screen "1. MAIN" 1280x800, template "Main_Template"
   on GenerateScreen: SetTag("animation_page", 1)
   Softkey "Softkey_F1" at 0,0 size 0x0
      on KeyDown: ActivateScreen("1. MAIN", 0)
   Softkey "Softkey_F2" at 0,0 size 0x0
      on KeyDown: ActivateScreen("2. VFD 2 - 5", 0)
   Softkey "Softkey_F3" at 0,0 size 0x0
      on KeyDown: ActivateScreen("3. VFD 6 - 9", 0)
   Softkey "Softkey_F4" at 0,0 size 0x0
      on KeyDown: ActivateScreen("4. VFD 10 - 13", 0)
   Softkey "Softkey_F5" at 0,0 size 0x0
      on KeyDown: ActivateScreen("5. VFD 14 - 17", 0)
   Softkey "Softkey_F6" at 0,0 size 0x0
      on KeyDown: ActivateScreen("6. VFD 18 - 21", 0)
   Softkey "Softkey_F7" at 0,0 size 0x0
      on KeyDown: ActivateScreen("7. VFD 22 - 23", 0)
   Softkey "Softkey_F8" at 0,0 size 0x0
      on KeyDown: ActivateScreen("8. ALARM", 0)
   Softkey "Softkey_F9" at 0,0 size 0x0
      on KeyDown: ActivateScreen("9. VFD PROFIBUS", 0)
   Softkey "Softkey_F10" at 0,0 size 0x0
      on KeyDown: ActivateScreen("10. SETTINGS", 0)
   TextField "Text field_33" at 632,247 size 105x42; Text 'Hz'
   TextField "Text field_1" at 0,64 size 331x50; Text 'ACTUAL MOTOR SPEED'
   Button "Button_1" at 0,721 size 160x79; TextOff 'MAIN'
      on Click: ActivateScreen("1. MAIN", 0)
      Appearance <- "animation_page"
   Button "Button_10" at 160,721 size 160x79; TextOff 'VFD 2 - 5'
      on Click: ActivateScreen("2. VFD 2 - 5", 0)
      Appearance <- "animation_page"
   Button "Button_11" at 320,721 size 160x79; TextOff 'VFD 6 - 9'
      on Click: ActivateScreen("3. VFD 6 - 9", 0)
      Appearance <- "animation_page"
   Button "Button_12" at 480,721 size 160x79; TextOff 'VFD 10 - 13'
      on Click: ActivateScreen("4. VFD 10 - 13", 0)
      Appearance <- "animation_page"
   Button "Button_13" at 640,721 size 160x79; TextOff 'VFD 14 - 17'
      on Click: ActivateScreen("5. VFD 14 - 17", 0)
      Appearance <- "animation_page"
   Button "Button_14" at 800,721 size 160x79; TextOff 'VFD 18 - 21'
      on Click: ActivateScreen("6. VFD 18 - 21", 0)
      Appearance <- "animation_page"
   Button "Button_15" at 960,721 size 160x79; TextOff 'VFD 22 - 23'
      on Click: ActivateScreen("7. VFD 22 - 23", 0)
      Appearance <- "animation_page"
   Button "Button_16" at 1120,721 size 160x79; TextOff 'Alarm'
      on Click: ActivateScreen("8. ALARM", 0)
      Appearance <- "animation_page"
   Group "Group" at 90,528 size 42x28
   Group "Group_1" at 57,540 size 42x28
   Group "Group_4" at 657,193 size 42x28
   Group "Group_5" at 3,194 size 42x28
   Group "Group_6" at 41,515 size 42x28
   Group "Group_15" at 926,512 size 42x28
   Group "Group_16" at 1063,535 size 42x28
   Group "Group_17" at 1008,534 size 42x28
   Group "Group_19" at 1058,421 size 42x28
   Group "Group_20" at 1103,421 size 42x28
   Group "Group_21" at 1165,505 size 42x28
   Group "Group_10" at 547,540 size 42x28
   Group "Group_9" at 510,515 size 42x28
   Group "Group_7" at 358,515 size 42x28
   Group "Group_8" at 396,540 size 42x28
   Group "Group_2" at 210,515 size 42x28
   Group "Group_3" at 252,540 size 42x28
   Group "Group_11" at 660,540 size 42x28
   Group "Group_12" at 797,502 size 42x28
   Group "Group_13" at 797,540 size 42x28
   Group "Group_14" at 853,530 size 42x28
   IOField "I/O field_17" at 633,252 size 60x33; FormatPattern 99.99
      ProcessValue <- "speedActual_address_18"
   TextField "Text field_24" at 22,247 size 105x42; Text 'Hz'
   IOField "I/O field_1" at 24,252 size 60x33; FormatPattern 99.99
      ProcessValue <- "speedActual_address_2"
   TextField "Text field_25" at 10,342 size 105x42; Text 'Hz'
   IOField "I/O field_2" at 12,347 size 60x33; FormatPattern 99.99
      ProcessValue <- "speedActual_address_3"
   Circle "Circle_34" at 693,170 size 28x28
      Appearance <- "Running_Motor Addres_23"
   Group "Group_18" at 1203,505 size 42x28
   Group "Group_22" at 1186,539 size 42x28
   Group "Group_23" at 11,162 size 42x28
   Group "Group_24" at 657,161 size 42x28
   TextField "Text field_29" at 33,653 size 105x42; Text 'Hz'
   IOField "I/O field_3" at 33,658 size 60x33; FormatPattern 99.99
      ProcessValue <- "speedActual_address_4"
   TextField "Text field_30" at 85,604 size 105x42; Text 'Hz'
   IOField "I/O field_4" at 87,609 size 60x33; FormatPattern 99.99
      ProcessValue <- "speedActual_address_5"
   TextField "Text field_31" at 177,653 size 105x42; Text 'Hz'
   IOField "I/O field_5" at 177,658 size 60x33; FormatPattern 99.99
      ProcessValue <- "speedActual_address_6"
   TextField "Text field_32" at 245,604 size 105x42; Text 'Hz'
   IOField "I/O field_6" at 247,609 size 60x33; FormatPattern 99.99
      ProcessValue <- "speedActual_address_7"
   TextField "Text field_34" at 322,653 size 105x42; Text 'Hz'
   IOField "I/O field_7" at 322,658 size 60x33; FormatPattern 99.99
      ProcessValue <- "speedActual_address_8"
   TextField "Text field_35" at 386,604 size 105x42; Text 'Hz'
   IOField "I/O field_8" at 388,609 size 60x33; FormatPattern 99.99
      ProcessValue <- "speedActual_address_9"
   TextField "Text field_36" at 467,653 size 105x42; Text 'Hz'
   IOField "I/O field_9" at 467,658 size 60x33; FormatPattern 99.99
      ProcessValue <- "speedActual_address_10"
   TextField "Text field_37" at 542,604 size 105x42; Text 'Hz'
   IOField "I/O field_10" at 544,609 size 60x33; FormatPattern 99.99
      ProcessValue <- "speedActual_address_11"
   TextField "Text field_38" at 611,653 size 105x42; Text 'Hz'
   IOField "I/O field_11" at 611,658 size 60x33; FormatPattern 99.99
      ProcessValue <- "speedActual_address_12"
   TextField "Text field_39" at 742,604 size 105x42; Text 'Hz'
   IOField "I/O field_12" at 744,609 size 60x33; FormatPattern 99.99
      ProcessValue <- "speedActual_address_13"
   TextField "Text field_40" at 756,653 size 105x42; Text 'Hz'
   IOField "I/O field_13" at 756,658 size 60x33; FormatPattern 99.99
      ProcessValue <- "speedActual_address_15"
   TextField "Text field_41" at 700,382 size 105x42; Text 'Hz'
   IOField "I/O field_14" at 702,387 size 60x33; FormatPattern 99.99
      ProcessValue <- "speedActual_address_14"
   TextField "Text field_42" at 901,653 size 105x42; Text 'Hz'
   IOField "I/O field_15" at 901,658 size 60x33; FormatPattern 99.99
      ProcessValue <- "speedActual_address_16"
   TextField "Text field_43" at 970,604 size 105x42; Text 'Hz'
   IOField "I/O field_16" at 972,609 size 60x33; FormatPattern 99.99
      ProcessValue <- "speedActual_address_17"
   TextField "Text field_44" at 1046,653 size 105x42; Text 'Hz'
   IOField "I/O field_18" at 1048,658 size 60x33; FormatPattern 99.99
      ProcessValue <- "speedActual_address_19"
   TextField "Text field_45" at 1150,604 size 105x42; Text 'Hz'
   IOField "I/O field_19" at 1152,609 size 60x33; FormatPattern 99.99
      ProcessValue <- "speedActual_address_22"
   TextField "Text field_46" at 1170,403 size 105x42; Text 'Hz'
   IOField "I/O field_20" at 1172,408 size 60x33; FormatPattern 99.99
      ProcessValue <- "speedActual_address_21"
   TextField "Text field_47" at 1170,325 size 105x42; Text 'Hz'
   IOField "I/O field_21" at 1172,330 size 60x33; FormatPattern 99.99
      ProcessValue <- "speedActual_address_20"
   TextField "Text field_48" at 1054,298 size 105x42; Text 'Hz'
   IOField "I/O field_22" at 1056,303 size 60x33; FormatPattern 99.99
      ProcessValue <- "speedActual_address_23"
   TextField "Text field_49" at 629,117 size 105x42; Text 'Hz'
   IOField "I/O field_23" at 631,122 size 60x33; FormatPattern 99.99
      ProcessValue <- "speedActual_address_23"
   TextField "Text field_50" at 13,117 size 105x42; Text 'Hz'
   IOField "I/O field_24" at 15,122 size 60x33; FormatPattern 99.99
      ProcessValue <- "speedActual_address_23"
   TextField "Text field_87" at 873,193 size 190x45; Text 'Rotary Moulder'
   Circle "Circle_10" at 883,201 size 29x29
      Appearance <- "Syncron_1"
   TextField "Text field_88" at 1071,141 size 190x45; Text 'Rotary Cutter'
   Circle "Circle_11" at 1081,149 size 29x29
      Appearance <- "Syncron_2"
   TextField "Text field_95" at 1071,193 size 190x45; Text 'Swivel Panner'
   Circle "Circle_12" at 1081,200 size 29x29
      Appearance <- "Syncron_3"
   TextField "Text field_51" at 873,141 size 190x45; Text 'SYNC MODE'
   TextField "Text field_52" at 42,320 size 42x25; Text '3'
   TextField "Text field_53" at 65,692 size 42x25; Text '4'
   TextField "Text field_54" at 117,582 size 42x25; Text '5'
   TextField "Text field_55" at 54,224 size 42x25; Text '2'
   TextField "Text field_56" at 635,224 size 42x25; Text '18'
   TextField "Text field_57" at 593,124 size 42x25; Text '23'
   TextField "Text field_58" at 121,124 size 42x25; Text '23'
   TextField "Text field_59" at 1086,276 size 42x25; Text '23'
   TextField "Text field_60" at 1173,582 size 42x25; Text '22'
   TextField "Text field_61" at 1202,300 size 42x25; Text '20'
   TextField "Text field_62" at 1202,376 size 42x25; Text '21'
   TextField "Text field_63" at 209,692 size 42x25; Text '6'
   TextField "Text field_64" at 277,582 size 42x25; Text '7'
   TextField "Text field_65" at 354,692 size 42x25; Text '8'
   TextField "Text field_66" at 418,582 size 42x25; Text '9'
   TextField "Text field_67" at 499,692 size 42x25; Text '10'
   TextField "Text field_68" at 574,582 size 42x25; Text '11'
   TextField "Text field_69" at 643,692 size 42x25; Text '12'
   TextField "Text field_70" at 788,692 size 42x25; Text '15'
   TextField "Text field_71" at 732,358 size 42x25; Text '14'
   TextField "Text field_72" at 990,582 size 42x25; Text '17'
   TextField "Text field_73" at 933,692 size 42x25; Text '16'
   TextField "Text field_74" at 1078,692 size 42x25; Text '19'
   TextField "Text field_75" at 774,582 size 42x25; Text '13'
   Button "Button_2" at 4,193 size 42x36; TextOff 'Text'
      on Click: ActivateScreen("2. VFD 2 - 5", 0)
   Button "Button_3" at 42,508 size 43x38; TextOff 'Text'
      on Click: ActivateScreen("2. VFD 2 - 5", 0)
   Button "Button_4" at 217,510 size 33x39; TextOff 'Text'
      on Click: ActivateScreen("3. VFD 6 - 9", 0)
   Button "Button_5" at 360,510 size 36x40; TextOff 'Text'
      on Click: ActivateScreen("3. VFD 6 - 9", 0)
   Button "Button_6" at 513,510 size 38x40; TextOff 'Text'
      on Click: ActivateScreen("4. VFD 10 - 13", 0)
   Button "Button_7" at 663,532 size 40x41; TextOff 'Text'
      on Click: ActivateScreen("4. VFD 10 - 13", 0)
   Button "Button_8" at 548,532 size 38x40; TextOff 'Text'
      on Click: ActivateScreen("4. VFD 10 - 13", 0)
   Button "Button_9" at 799,532 size 40x41; TextOff 'Text'
      on Click: ActivateScreen("4. VFD 10 - 13", 0)
   Button "Button_17" at 855,524 size 40x41; TextOff 'Text'
      on Click: ActivateScreen("5. VFD 14 - 17", 0)
   Button "Button_18" at 799,492 size 40x41; TextOff 'Text'
      on Click: ActivateScreen("5. VFD 14 - 17", 0)
   Button "Button_19" at 927,508 size 40x41; TextOff 'Text'
      on Click: ActivateScreen("5. VFD 14 - 17", 0)
   Button "Button_20" at 1007,524 size 40x41; TextOff 'Text'
      on Click: ActivateScreen("5. VFD 14 - 17", 0)
   Button "Button_21" at 1064,526 size 40x41; TextOff 'Text'
      on Click: ActivateScreen("6. VFD 18 - 21", 0)
   Button "Button_22" at 1187,539 size 40x31; TextOff 'Text'
      on Click: ActivateScreen("7. VFD 22 - 23", 0)
   Button "Button_23" at 1165,497 size 82x41; TextOff 'Text'
      on Click: ActivateScreen("6. VFD 18 - 21", 0)
   Button "Button_24" at 1060,414 size 40x39; TextOff 'Text'
      on Click: ActivateScreen("7. VFD 22 - 23", 0)
   Button "Button_25" at 1105,414 size 40x39; TextOff 'Text'
      on Click: ActivateScreen("7. VFD 22 - 23", 0)
   Button "Button_26" at 659,156 size 40x39; TextOff 'Text'
      on Click: ActivateScreen("7. VFD 22 - 23", 0)
   Button "Button_27" at 13,156 size 40x39; TextOff 'Text'
      on Click: ActivateScreen("7. VFD 22 - 23", 0)
   Button "Button_28" at 659,190 size 40x41; TextOff 'Text'
      on Click: ActivateScreen("6. VFD 18 - 21", 0)
   Button "Button_29" at 400,533 size 36x40; TextOff 'Text'
      on Click: ActivateScreen("3. VFD 6 - 9", 0)
   Button "Button_30" at 257,534 size 33x39; TextOff 'Text'
      on Click: ActivateScreen("3. VFD 6 - 9", 0)
   Button "Button_31" at 58,532 size 43x38; TextOff 'Text'
      on Click: ActivateScreen("2. VFD 2 - 5", 0)
   Button "Button_32" at 90,524 size 43x38; TextOff 'Text'
      on Click: ActivateScreen("2. VFD 2 - 5", 0)
   Circle "Circle_2" at 97,528 size 28x28
      Appearance <- "Running_Motor Addres_5"
   TextField "Text field_2" at 90,530 size 42x25; Text 'M'
   Circle "Circle_23" at 64,540 size 28x28
      Appearance <- "Running_Motor Addres_4"
   TextField "Text field_3" at 57,542 size 42x25; Text 'M'
   Circle "Circle_6" at 664,193 size 28x28
      Appearance <- "Running_Motor Addres_18"
   TextField "Text field_6" at 657,195 size 42x25; Text 'M'
   Circle "Circle_22" at 10,194 size 28x28
      Appearance <- "Running_Motor Addres_2"
   TextField "Text field_7" at 3,196 size 42x25; Text 'M'
   Circle "Circle_5" at 48,515 size 28x28
      Appearance <- "Running_Motor Addres_3"
   TextField "Text field_8" at 41,517 size 42x25; Text 'M'
   Circle "Circle_31" at 933,512 size 28x28
      Appearance <- "Running_Motor Addres_16"
   TextField "Text field_17" at 926,514 size 42x25; Text 'M'
   Circle "Circle_32" at 1070,535 size 28x28
      Appearance <- "Running_Motor Addres_19"
   TextField "Text field_18" at 1063,537 size 42x25; Text 'M'
   Circle "Circle_33" at 1015,534 size 28x28
      Appearance <- "Running_Motor Addres_17"
   TextField "Text field_19" at 1008,536 size 42x25; Text 'M'
   Circle "Circle_35" at 1065,421 size 28x28
      Appearance <- "Running_Motor Addres_23"
   TextField "Text field_21" at 1058,423 size 42x25; Text 'M'
   Circle "Circle_36" at 1110,421 size 28x28
      Appearance <- "Running_Motor Addres_23"
   TextField "Text field_22" at 1103,423 size 42x25; Text 'M'
   Circle "Circle_37" at 1172,505 size 28x28
      Appearance <- "Running_Motor Addres_20"
   TextField "Text field_23" at 1165,507 size 42x25; Text 'M'
   Circle "Circle_26" at 554,540 size 28x28
      Appearance <- "Running_Motor Addres_11"
   TextField "Text field_12" at 547,542 size 42x25; Text 'M'
   Circle "Circle_25" at 517,515 size 28x28
      Appearance <- "Running_Motor Addres_10"
   TextField "Text field_11" at 510,517 size 42x25; Text 'M'
   Circle "Circle_21" at 365,515 size 28x28
      Appearance <- "Running_Motor Addres_8"
   TextField "Text field_9" at 358,517 size 42x25; Text 'M'
   Circle "Circle_24" at 403,540 size 28x28
      Appearance <- "Running_Motor Addres_9"
   TextField "Text field_10" at 396,542 size 42x25; Text 'M'
   Circle "Circle_1" at 217,515 size 28x28
      Appearance <- "Running_Motor Addres_6"
   TextField "Text field_4" at 210,517 size 42x25; Text 'M'
   Circle "Circle_7" at 259,540 size 28x28
      Appearance <- "Running_Motor Addres_7"
   TextField "Text field_5" at 252,542 size 42x25; Text 'M'
   Circle "Circle_27" at 667,540 size 28x28
      Appearance <- "Running_Motor Addres_12"
   TextField "Text field_13" at 660,542 size 42x25; Text 'M'
   Circle "Circle_28" at 804,502 size 28x28
      Appearance <- "Running_Motor Addres_14"
   TextField "Text field_14" at 797,504 size 42x25; Text 'M'
   Circle "Circle_29" at 804,540 size 28x28
      Appearance <- "Running_Motor Addres_13"
   TextField "Text field_15" at 797,542 size 42x25; Text 'M'
   Circle "Circle_30" at 860,530 size 28x28
      Appearance <- "Running_Motor Addres_15"
   TextField "Text field_16" at 853,532 size 42x25; Text 'M'
   Circle "Circle_3" at 1210,505 size 28x28
      Appearance <- "Running_Motor Addres_21"
   TextField "Text field_20" at 1203,507 size 42x25; Text 'M'
   Circle "Circle_4" at 1193,539 size 28x28
      Appearance <- "Running_Motor Addres_22"
   TextField "Text field_26" at 1186,541 size 42x25; Text 'M'
   Circle "Circle_8" at 18,162 size 28x28
      Appearance <- "Running_Motor Addres_23"
   TextField "Text field_27" at 11,164 size 42x25; Text 'M'
   Circle "Circle_9" at 664,161 size 28x28
      Appearance <- "Running_Motor Addres_23"
   TextField "Text field_28" at 657,163 size 42x25; Text 'M'

screen "8. ALARM" 1280x800, template "Main_Template"
   on GenerateScreen: SetTag("animation_page", 8)
   Softkey "Softkey_F1" at 0,0 size 0x0
      on KeyDown: ActivateScreen("1. MAIN", 0)
   Softkey "Softkey_F2" at 0,0 size 0x0
      on KeyDown: ActivateScreen("2. VFD 2 - 5", 0)
   Softkey "Softkey_F3" at 0,0 size 0x0
      on KeyDown: ActivateScreen("3. VFD 6 - 9", 0)
   Softkey "Softkey_F4" at 0,0 size 0x0
      on KeyDown: ActivateScreen("4. VFD 10 - 13", 0)
   Softkey "Softkey_F5" at 0,0 size 0x0
      on KeyDown: ActivateScreen("5. VFD 14 - 17", 0)
   Softkey "Softkey_F6" at 0,0 size 0x0
      on KeyDown: ActivateScreen("6. VFD 18 - 21", 0)
   Softkey "Softkey_F7" at 0,0 size 0x0
      on KeyDown: ActivateScreen("7. VFD 22 - 23", 0)
   Softkey "Softkey_F8" at 0,0 size 0x0
      on KeyDown: ActivateScreen("8. ALARM", 0)
   Softkey "Softkey_F9" at 0,0 size 0x0
      on KeyDown: ActivateScreen("9. VFD PROFIBUS", 0)
   AlarmView "Alarm view_1" at 38,140 size 1199x553
   TextField "Text field_38" at 0,64 size 331x50; Text 'ALARMS'
   Button "Button_1" at 0,721 size 160x79; TextOff 'MAIN'
      on Click: ActivateScreen("1. MAIN", 0)
      Appearance <- "animation_page"
   Button "Button_10" at 160,721 size 160x79; TextOff 'VFD 2 - 5'
      on Click: ActivateScreen("2. VFD 2 - 5", 0)
      Appearance <- "animation_page"
   Button "Button_11" at 320,721 size 160x79; TextOff 'VFD 6 - 9'
      on Click: ActivateScreen("3. VFD 6 - 9", 0)
      Appearance <- "animation_page"
   Button "Button_12" at 480,721 size 160x79; TextOff 'VFD 10 - 13'
      on Click: ActivateScreen("4. VFD 10 - 13", 0)
      Appearance <- "animation_page"
   Button "Button_13" at 640,721 size 160x79; TextOff 'VFD 14 - 17'
      on Click: ActivateScreen("5. VFD 14 - 17", 0)
      Appearance <- "animation_page"
   Button "Button_14" at 800,721 size 160x79; TextOff 'VFD 18 - 21'
      on Click: ActivateScreen("6. VFD 18 - 21", 0)
      Appearance <- "animation_page"
   Button "Button_15" at 960,721 size 160x79; TextOff 'VFD 22 - 23'
      on Click: ActivateScreen("7. VFD 22 - 23", 0)
      Appearance <- "animation_page"
   Button "Button_16" at 1120,721 size 160x79; TextOff 'Alarm'
      on Click: ActivateScreen("8. ALARM", 0)
      Appearance <- "animation_page"
   Softkey "Softkey_F10" at 0,0 size 0x0
      on KeyDown: ActivateScreen("10. SETTINGS", 0)

screen "11. DIAG" 1280x800, template "Main_Template"
   on GenerateScreen: function_fa202464("System diagnostics view_1"); SetTag("animation_page", 0)
   SysDiagControl "System diagnostics view_1" at 35,130 size 1206x565
   TextField "Text field_38" at 0,64 size 331x50; Text 'SYSTEM DIAGNOSTIC'
   Button "Button_1" at 0,721 size 160x79; TextOff 'MAIN'
      on Click: ActivateScreen("1. MAIN", 0)
   Button "Button_10" at 160,721 size 160x79; TextOff 'VFD 2 - 5'
      on Click: ActivateScreen("2. VFD 2 - 5", 0)
   Button "Button_11" at 320,721 size 160x79; TextOff 'VFD 6 - 9'
      on Click: ActivateScreen("3. VFD 6 - 9", 0)
   Button "Button_12" at 480,721 size 160x79; TextOff 'VFD 10 - 13'
      on Click: ActivateScreen("4. VFD 10 - 13", 0)
   Button "Button_13" at 640,721 size 160x79; TextOff 'VFD 14 - 17'
      on Click: ActivateScreen("5. VFD 14 - 17", 0)
   Button "Button_14" at 800,721 size 160x79; TextOff 'VFD 18 - 21'
      on Click: ActivateScreen("6. VFD 18 - 21", 0)
   Button "Button_15" at 960,721 size 160x79; TextOff 'VFD 22 - 23'
      on Click: ActivateScreen("7. VFD 22 - 23", 0)
   Button "Button_16" at 1120,721 size 160x79; TextOff 'Alarm'
      on Click: ActivateScreen("8. ALARM", 0)
   Softkey "Softkey_F1" at 0,0 size 0x0
      on KeyDown: ActivateScreen("1. MAIN", 0)
   Softkey "Softkey_F2" at 0,0 size 0x0
      on KeyDown: ActivateScreen("2. VFD 2 - 5", 0)
   Softkey "Softkey_F3" at 0,0 size 0x0
      on KeyDown: ActivateScreen("3. VFD 6 - 9", 0)
   Softkey "Softkey_F4" at 0,0 size 0x0
      on KeyDown: ActivateScreen("4. VFD 10 - 13", 0)
   Softkey "Softkey_F5" at 0,0 size 0x0
      on KeyDown: ActivateScreen("5. VFD 14 - 17", 0)
   Softkey "Softkey_F6" at 0,0 size 0x0
      on KeyDown: ActivateScreen("6. VFD 18 - 21", 0)
   Softkey "Softkey_F7" at 0,0 size 0x0
      on KeyDown: ActivateScreen("7. VFD 22 - 23", 0)
   Softkey "Softkey_F8" at 0,0 size 0x0
      on KeyDown: ActivateScreen("8. ALARM", 0)
   Softkey "Softkey_F9" at 0,0 size 0x0
      on KeyDown: ActivateScreen("9. VFD PROFIBUS", 0)
   Softkey "Softkey_F10" at 0,0 size 0x0
      on KeyDown: ActivateScreen("10. SETTINGS", 0)

screen "10. SETTINGS" 1280x800, template "Main_Template"
   on GenerateScreen: SetTag("animation_page", 0)
   GraphicView "Graphic view_4" at 11,688 size 244x98; Picture "Graphic_9"
   Button "Button_1" at 11,688 size 244x98; TextOff 'Text'
      on Click: StopRuntime(0)
   TextField "Text field_2" at 342,188 size 247x54; Text 'Date Time Setting'
   DateTimeField "Date/time field_1" at 534,264 size 604x89; Authorization "User administration"
   Button "Button_2" at 11,123 size 244x98; TextOff 'Overview / DI / DO VIEW'
      on Click: ActivateScreen("12. DI/DO", 0)
      Appearance <- "animation_page"
   Button "Button_6" at 11,264 size 244x98; TextOff 'Alarm'
      on Click: SetTag("animation_page", 6); ActivateScreen("8. ALARM", 0)
      Appearance <- "animation_page"
   Button "Button_3" at 11,405 size 244x98; TextOff 'Calibrate Screen'
      on Click: function_bc3e350c()
      Appearance <- "animation_page"
   Button "Button_4" at 11,546 size 244x98; TextOff 'Clean Screen'
      on Click: function_be740847(30)
      Appearance <- "animation_page"
   TextField "Text field_38" at 0,64 size 331x50; Text 'SETINGS'
   Button "Button_8" at 908,688 size 244x98; TextOff 'Communication Overview'
      on Click: ActivateScreen("9. VFD PROFIBUS", 0)
      Appearance <- "animation_page"
   DateTimeField "Date/time field_2" at 534,408 size 604x89
   TextField "Text field_1" at 368,290 size 85x37; Text 'DATE'
   TextField "Text field_3" at 368,434 size 76x37; Text 'TIME'
   Softkey "Softkey_F1" at 0,0 size 0x0
      on KeyDown: ActivateScreen("1. MAIN", 0)
   Softkey "Softkey_F2" at 0,0 size 0x0
      on KeyDown: ActivateScreen("2. VFD 2 - 5", 0)
   Softkey "Softkey_F3" at 0,0 size 0x0
      on KeyDown: ActivateScreen("3. VFD 6 - 9", 0)
   Softkey "Softkey_F4" at 0,0 size 0x0
      on KeyDown: ActivateScreen("4. VFD 10 - 13", 0)
   Softkey "Softkey_F5" at 0,0 size 0x0
      on KeyDown: ActivateScreen("5. VFD 14 - 17", 0)
   Softkey "Softkey_F6" at 0,0 size 0x0
      on KeyDown: ActivateScreen("6. VFD 18 - 21", 0)
   Softkey "Softkey_F7" at 0,0 size 0x0
      on KeyDown: ActivateScreen("7. VFD 22 - 23", 0)
   Softkey "Softkey_F8" at 0,0 size 0x0
      on KeyDown: ActivateScreen("8. ALARM", 0)
   Softkey "Softkey_F9" at 0,0 size 0x0
      on KeyDown: ActivateScreen("9. VFD PROFIBUS", 0)
   Softkey "Softkey_F10" at 0,0 size 0x0
      on KeyDown: ActivateScreen("10. SETTINGS", 0)

screen "9. VFD PROFIBUS" 1280x800, template "Main_Template"
   on GenerateScreen: SetTag("animation_page", 0)
   TextField "Text field_1" at 116,456 size 30x30; Text '2'
      Appearance <- "Address_2"
   TextField "Text field_2" at 116,665 size 30x30; Text '13'
      Appearance <- "Address_13"
   TextField "Text field_3" at 220,456 size 30x30; Text '3'
      Appearance <- "Address_3"
   TextField "Text field_4" at 324,456 size 30x30; Text '4'
      Appearance <- "Address_4"
   TextField "Text field_5" at 428,456 size 30x30; Text '5'
      Appearance <- "Address_5"
   TextField "Text field_6" at 532,456 size 30x30; Text '6'
      Appearance <- "Address_6"
   TextField "Text field_7" at 636,456 size 30x30; Text '7'
      Appearance <- "Address_7"
   TextField "Text field_8" at 740,456 size 30x30; Text '8'
      Appearance <- "Address_8"
   TextField "Text field_9" at 844,456 size 30x30; Text '9'
      Appearance <- "Address_9"
   TextField "Text field_10" at 948,456 size 30x30; Text '10'
      Appearance <- "Address_10"
   TextField "Text field_11" at 1052,456 size 30x30; Text '11'
      Appearance <- "Address_11"
   TextField "Text field_12" at 1156,456 size 30x30; Text '12'
      Appearance <- "Address_12"
   TextField "Text field_13" at 220,665 size 30x30; Text '14'
      Appearance <- "Address_14"
   TextField "Text field_14" at 324,665 size 30x30; Text '15'
      Appearance <- "Address_15"
   TextField "Text field_15" at 428,665 size 30x30; Text '16'
      Appearance <- "Address_16"
   TextField "Text field_16" at 532,665 size 30x30; Text '17'
      Appearance <- "Address_17"
   TextField "Text field_17" at 636,665 size 30x30; Text '18'
      Appearance <- "Address_18"
   TextField "Text field_18" at 740,665 size 30x30; Text '19'
      Appearance <- "Address_19"
   TextField "Text field_19" at 844,665 size 30x30; Text '20'
      Appearance <- "Address_20"
   TextField "Text field_20" at 948,665 size 30x30; Text '21'
      Appearance <- "Address_21"
   TextField "Text field_21" at 1052,665 size 30x30; Text '22'
      Appearance <- "Address_22"
   TextField "Text field_22" at 1156,665 size 30x30; Text '23'
      Appearance <- "Address_23"
   TextField "Text field_38" at 0,64 size 331x50; Text 'COMMUNICATION'
   TextField "Text field_23" at 1063,145 size 74x25; Text 'PLC'
   TextField "Text field_24" at 438,145 size 74x25; Text 'HMI'
   TextField "Text field_25" at 75,314 size 71x25; Text 'VFD 2'
      Appearance <- "Running_Motor Addres_2"
   TextField "Text field_26" at 179,314 size 71x25; Text 'VFD 3'
      Appearance <- "Running_Motor Addres_3"
   TextField "Text field_27" at 283,314 size 71x25; Text 'VFD 4'
      Appearance <- "Running_Motor Addres_4"
   TextField "Text field_28" at 387,314 size 71x25; Text 'VFD 5'
      Appearance <- "Running_Motor Addres_5"
   TextField "Text field_29" at 491,314 size 71x25; Text 'VFD 6'
      Appearance <- "Running_Motor Addres_6"
   TextField "Text field_30" at 595,314 size 71x25; Text 'VFD 7'
      Appearance <- "Running_Motor Addres_7"
   TextField "Text field_31" at 699,314 size 71x25; Text 'VFD 8'
      Appearance <- "Running_Motor Addres_8"
   TextField "Text field_32" at 803,314 size 71x25; Text 'VFD 9'
      Appearance <- "Running_Motor Addres_9"
   TextField "Text field_33" at 907,314 size 71x25; Text 'VFD 10'
      Appearance <- "Running_Motor Addres_10"
   TextField "Text field_34" at 1011,314 size 71x25; Text 'VFD 11'
      Appearance <- "Running_Motor Addres_11"
   TextField "Text field_35" at 1115,314 size 71x25; Text 'VFD 12'
      Appearance <- "Running_Motor Addres_12"
   TextField "Text field_36" at 75,522 size 71x25; Text 'VFD 13'
      Appearance <- "Running_Motor Addres_13"
   TextField "Text field_37" at 179,522 size 71x25; Text 'VFD 14'
      Appearance <- "Running_Motor Addres_14"
   TextField "Text field_39" at 283,522 size 71x25; Text 'VFD 15'
      Appearance <- "Running_Motor Addres_15"
   TextField "Text field_40" at 387,522 size 71x25; Text 'VFD 16'
      Appearance <- "Running_Motor Addres_16"
   TextField "Text field_41" at 491,522 size 71x25; Text 'VFD 17'
      Appearance <- "Running_Motor Addres_17"
   TextField "Text field_42" at 595,522 size 71x25; Text 'VFD 18'
      Appearance <- "Running_Motor Addres_18"
   TextField "Text field_43" at 699,522 size 71x25; Text 'VFD 19'
      Appearance <- "Running_Motor Addres_19"
   TextField "Text field_44" at 803,522 size 71x25; Text 'VFD 20'
      Appearance <- "Running_Motor Addres_20"
   TextField "Text field_45" at 907,522 size 71x25; Text 'VFD 21'
      Appearance <- "Running_Motor Addres_21"
   TextField "Text field_46" at 1011,522 size 71x25; Text 'VFD 22'
      Appearance <- "Running_Motor Addres_22"
   TextField "Text field_47" at 1115,522 size 71x25; Text 'VFD 23'
      Appearance <- "Running_Motor Addres_23"
   TextField "Text field_48" at 306,165 size 82x25; Text 'KTP1200'
   IOField "I/O field_2" at 185,354 size 59x27; FormatPattern 99.99
      ProcessValue <- "speedActual_address_3"
   IOField "I/O field_3" at 289,354 size 59x27; FormatPattern 99.99
      ProcessValue <- "speedActual_address_4"
   IOField "I/O field_4" at 393,354 size 59x27; FormatPattern 99.99
      ProcessValue <- "speedActual_address_5"
   IOField "I/O field_5" at 497,354 size 59x27; FormatPattern 99.99
      ProcessValue <- "speedActual_address_6"
   IOField "I/O field_6" at 601,354 size 59x27; FormatPattern 99.99
      ProcessValue <- "speedActual_address_7"
   IOField "I/O field_7" at 705,354 size 59x27; FormatPattern 99.99
      ProcessValue <- "speedActual_address_8"
   IOField "I/O field_8" at 809,354 size 59x27; FormatPattern 99.99
      ProcessValue <- "speedActual_address_9"
   IOField "I/O field_9" at 913,354 size 59x27; FormatPattern 99.99
      ProcessValue <- "speedActual_address_10"
   IOField "I/O field_10" at 1017,354 size 59x27; FormatPattern 99.99
      ProcessValue <- "speedActual_address_11"
   IOField "I/O field_11" at 1121,354 size 59x27; FormatPattern 99.99
      ProcessValue <- "speedActual_address_12"
   IOField "I/O field_12" at 81,562 size 59x27; FormatPattern 99.99
      ProcessValue <- "speedActual_address_13"
   IOField "I/O field_13" at 185,562 size 59x27; FormatPattern 99.99
      ProcessValue <- "speedActual_address_14"
   IOField "I/O field_14" at 289,562 size 59x27; FormatPattern 99.99
      ProcessValue <- "speedActual_address_15"
   IOField "I/O field_15" at 393,562 size 59x27; FormatPattern 99.99
      ProcessValue <- "speedActual_address_16"
   IOField "I/O field_16" at 497,562 size 59x27; FormatPattern 99.99
      ProcessValue <- "speedActual_address_17"
   IOField "I/O field_17" at 601,562 size 59x27; FormatPattern 99.99
      ProcessValue <- "speedActual_address_18"
   IOField "I/O field_18" at 705,562 size 59x27; FormatPattern 99.99
      ProcessValue <- "speedActual_address_19"
   IOField "I/O field_19" at 809,562 size 59x27; FormatPattern 99.99
      ProcessValue <- "speedActual_address_20"
   IOField "I/O field_20" at 913,562 size 59x27; FormatPattern 99.99
      ProcessValue <- "speedActual_address_21"
   IOField "I/O field_21" at 1017,562 size 59x27; FormatPattern 99.99
      ProcessValue <- "speedActual_address_22"
   IOField "I/O field_22" at 1121,562 size 59x27; FormatPattern 99.99
      ProcessValue <- "speedActual_address_23"
   IOField "I/O field_1" at 81,354 size 59x27; FormatPattern 99.99
      ProcessValue <- "speedActual_address_2"
   Button "Button_1" at 820,122 size 239x120; TextOff '12.DI/DO'
      on Click: ActivateScreen("12. DI/DO", 0)
   Softkey "Softkey_F1" at 0,0 size 0x0
      on KeyDown: ActivateScreen("1. MAIN", 0)
   Softkey "Softkey_F2" at 0,0 size 0x0
      on KeyDown: ActivateScreen("2. VFD 2 - 5", 0)
   Softkey "Softkey_F3" at 0,0 size 0x0
      on KeyDown: ActivateScreen("3. VFD 6 - 9", 0)
   Softkey "Softkey_F4" at 0,0 size 0x0
      on KeyDown: ActivateScreen("4. VFD 10 - 13", 0)
   Softkey "Softkey_F5" at 0,0 size 0x0
      on KeyDown: ActivateScreen("5. VFD 14 - 17", 0)
   Softkey "Softkey_F6" at 0,0 size 0x0
      on KeyDown: ActivateScreen("6. VFD 18 - 21", 0)
   Softkey "Softkey_F7" at 0,0 size 0x0
      on KeyDown: ActivateScreen("7. VFD 22 - 23", 0)
   Softkey "Softkey_F8" at 0,0 size 0x0
      on KeyDown: ActivateScreen("8. ALARM", 0)
   Softkey "Softkey_F9" at 0,0 size 0x0
      on KeyDown: ActivateScreen("9. VFD PROFIBUS", 0)
   Softkey "Softkey_F10" at 0,0 size 0x0
      on KeyDown: ActivateScreen("10. SETTINGS", 0)

Template "Main_Template" 1280x800
   TextField "Template_Text field_1" at 10,14 size 388x39; Text 'FORMING LINE MACHINE'
   TextField "Template_Text field_2" at 986,64 size 294x50; Text 'Rotary Moulder Mode'
      Visibility <- "Rotary_Moulder"
   TextField "Template_Text field_3" at 986,64 size 294x50; Text 'Rotary Cutter Mode'
      Visibility <- "Rotary_Cutting"
   GraphicView "Template_Graphic view_1" at 398,0 size 136x64; Picture "biru"
   DateTimeField "Template_Date/time field_1" at 986,18 size 272x30
   GraphicView "Template_Graphic view_2" at 894,4 size 72x59; Picture "emc"
      Visibility <- "EMERGENCY"
      Appearance <- "EMERGENCY"

screen "2. VFD 2 - 5" 1280x800, template "Main_Template"
   on GenerateScreen: SetTag("animation_page", 2)
   Bar "Bar_1" at 206,213 size 88x440; MinimumValue 0; MaximumValue 50
      ProcessValue <- "speedActual_address_2"
   Button "Button_7" at 35,514 size 150x62; TextOff '+'
      on Press: function_b14e0dd5("increaseSpeed_address_2", 0)
      Appearance <- "statusIncrease_address_2"
   Button "Button_8" at 35,591 size 150x62; TextOff '-'
      on Press: function_b14e0dd5("decreaseSpeed_address_2", 0)
      Appearance <- "statusDecrease_address_2"
   TextField "Text field_20" at 35,428 size 150x62; Text 'Hz'
   IOField "I/O field_1" at 37,430 size 98x57; FormatPattern 99.99
      ProcessValue <- "speedActual_address_2"
   TextField "Text field_14" at 28,133 size 207x62; Text 'Conveyor of Metal Detector'
   TextField "Text field_26" at 35,228 size 150x62; Text 'Hz'
   TextField "Text field_32" at 35,328 size 150x62; Text '-'
   IOField "I/O field_2" at 39,231 size 98x57; FormatPattern 99.99
      ProcessValue <- "speedReff_singleSync_address_2"
   TextField "Text field_1" at 35,400 size 115x27; Text 'Actual Speed'
   TextField "Text field_2" at 35,302 size 144x27; Text 'Reff Speed Sync'
   TextField "Text field_3" at 35,200 size 155x27; Text 'Reff Speed Single'
   TextField "Text field_4" at 36,661 size 149x45; Text 'VFD 2'
      Appearance <- "Running_Motor Addres_2"
   Bar "Bar_2" at 518,213 size 88x440; MinimumValue 0; MaximumValue 50
      ProcessValue <- "speedActual_address_3"
   Button "Button_2" at 347,514 size 150x62; TextOff '+'
      on Press: function_b14e0dd5("increaseSpeed_address_3", 0)
      Appearance <- "statusIncrease_address_3"
   Button "Button_3" at 347,591 size 150x62; TextOff '-'
      on Press: function_b14e0dd5("decreaseSpeed_address_3", 0)
      Appearance <- "statusDecrease_address_3"
   TextField "Text field_5" at 347,428 size 150x62; Text 'Hz'
   IOField "I/O field_3" at 349,430 size 98x57; FormatPattern 99.99
      ProcessValue <- "speedActual_address_3"
   TextField "Text field_6" at 340,133 size 207x62; Text 'Gauge Roll 2nd Set'
   TextField "Text field_7" at 347,228 size 150x62; Text 'Hz'
   TextField "Text field_8" at 347,328 size 150x62; Text 'Hz'
   IOField "I/O field_4" at 351,231 size 98x57; FormatPattern 99.99
      ProcessValue <- "speedReff_singleSync_address_3"
   TextField "Text field_9" at 347,400 size 115x27; Text 'Actual Speed'
   TextField "Text field_10" at 347,302 size 144x27; Text 'Reff Speed Sync'
   TextField "Text field_11" at 347,200 size 155x27; Text 'Reff Speed Single'
   TextField "Text field_12" at 348,661 size 149x45; Text 'VFD 3'
      Appearance <- "Running_Motor Addres_3"
   Bar "Bar_3" at 830,213 size 88x440; MinimumValue 0; MaximumValue 50
      ProcessValue <- "speedActual_address_4"
   Button "Button_4" at 659,514 size 150x62; TextOff '+'
      on Press: function_b14e0dd5("increaseSpeed_address_4", 0)
      Appearance <- "statusIncrease_address_4"
   Button "Button_5" at 659,591 size 150x62; TextOff '-'
      on Press: function_b14e0dd5("decreaseSpeed_address_4", 0)
      Appearance <- "statusDecrease_address_4"
   TextField "Text field_13" at 659,428 size 150x62; Text 'Hz'
   IOField "I/O field_5" at 661,430 size 98x57; FormatPattern 99.99
      ProcessValue <- "speedActual_address_4"
   TextField "Text field_15" at 652,133 size 207x62; Text 'Gauge Roll 1st Set'
   TextField "Text field_16" at 659,228 size 150x62; Text 'Hz'
   TextField "Text field_17" at 659,328 size 150x62; Text 'Hz'
   IOField "I/O field_6" at 663,231 size 98x57; FormatPattern 99.99
      ProcessValue <- "speedReff_singleSync_address_4"
   TextField "Text field_18" at 659,400 size 115x27; Text 'Actual Speed'
   TextField "Text field_19" at 659,302 size 144x27; Text 'Reff Speed Sync'
   TextField "Text field_21" at 659,200 size 155x27; Text 'Reff Speed Single'
   TextField "Text field_22" at 660,661 size 149x45; Text 'VFD 4'
      Appearance <- "Running_Motor Addres_4"
   Bar "Bar_4" at 1142,213 size 88x440; MinimumValue 0; MaximumValue 50
      ProcessValue <- "speedActual_address_5"
   Button "Button_6" at 971,514 size 150x62; TextOff '+'
      on Press: function_b14e0dd5("increaseSpeed_address_5", 0)
      Appearance <- "statusIncrease_address_5"
   Button "Button_9" at 971,591 size 150x62; TextOff '-'
      on Press: function_b14e0dd5("decreaseSpeed_address_5", 0)
      Appearance <- "statusDecrease_address_5"
   TextField "Text field_23" at 971,428 size 150x62; Text 'Hz'
   IOField "I/O field_7" at 973,430 size 98x57; FormatPattern 99.99
      ProcessValue <- "speedActual_address_5"
   TextField "Text field_24" at 964,133 size 207x62; Text 'Passing Conveyor 3-Roll Sheeter'
   TextField "Text field_25" at 971,228 size 150x62; Text 'Hz'
   TextField "Text field_27" at 971,328 size 150x62; Text 'Hz'
   IOField "I/O field_8" at 975,231 size 98x57; FormatPattern 99.99
      ProcessValue <- "speedReff_singleSync_address_5"
   TextField "Text field_28" at 971,400 size 115x27; Text 'Actual Speed'
   TextField "Text field_29" at 971,302 size 144x27; Text 'Reff Speed Sync'
   TextField "Text field_30" at 971,200 size 155x27; Text 'Reff Speed Single'
   TextField "Text field_31" at 972,661 size 149x45; Text 'VFD 5'
      Appearance <- "Running_Motor Addres_5"
   IOField "I/O field_14" at 349,330 size 98x57; FormatPattern 99.99
      ProcessValue <- "speedReff_NOT_singleSync_address_3"
   IOField "I/O field_9" at 661,330 size 98x57; FormatPattern 99.99
      ProcessValue <- "speedReff_NOT_singleSync_address_4"
   IOField "I/O field_10" at 973,330 size 98x57; FormatPattern 99.99
      ProcessValue <- "speedReff_NOT_singleSync_address_5"
   SymbolicIOField "Symbolic I/O field_2" at 550,133 size 77x62; TextOn '1'; TextOff '0'; TextList "Mode_Syncron"
      Appearance <- "Syncron_2"
      ProcessValue <- "Syncron_2"
   SymbolicIOField "Symbolic I/O field_3" at 862,133 size 77x62; TextOn '1'; TextOff '0'; TextList "Mode_Syncron"
      Appearance <- "Syncron_2"
      ProcessValue <- "Syncron_2"
   SymbolicIOField "Symbolic I/O field_4" at 1174,133 size 77x62; TextOn '1'; TextOff '0'; TextList "Mode_Syncron"
      Appearance <- "Syncron_2"
      ProcessValue <- "Syncron_2"
   TextField "Text field_33" at 238,133 size 76x62; Text 'Single'
   Button "Button_1" at 0,721 size 160x79; TextOff 'MAIN'
      on Click: ActivateScreen("1. MAIN", 0)
      Appearance <- "animation_page"
   Button "Button_10" at 160,721 size 160x79; TextOff 'VFD 2 - 5'
      on Click: ActivateScreen("2. VFD 2 - 5", 0)
      Appearance <- "animation_page"
   Button "Button_11" at 320,721 size 160x79; TextOff 'VFD 6 - 9'
      on Click: ActivateScreen("3. VFD 6 - 9", 0)
      Appearance <- "animation_page"
   Button "Button_12" at 480,721 size 160x79; TextOff 'VFD 10 - 13'
      on Click: ActivateScreen("4. VFD 10 - 13", 0)
      Appearance <- "animation_page"
   Button "Button_13" at 640,721 size 160x79; TextOff 'VFD 14 - 17'
      on Click: ActivateScreen("5. VFD 14 - 17", 0)
      Appearance <- "animation_page"
   Button "Button_14" at 800,721 size 160x79; TextOff 'VFD 18 - 21'
      on Click: ActivateScreen("6. VFD 18 - 21", 0)
      Appearance <- "animation_page"
   Button "Button_15" at 960,721 size 160x79; TextOff 'VFD 22 - 23'
      on Click: ActivateScreen("7. VFD 22 - 23", 0)
      Appearance <- "animation_page"
   Button "Button_16" at 1120,721 size 160x79; TextOff 'Alarm'
      on Click: ActivateScreen("8. ALARM", 0)
      Appearance <- "animation_page"
   TextField "Text field_34" at 0,64 size 331x50; Text 'MOTOR CONTROL SPEED'
   Softkey "Softkey_F1" at 0,0 size 0x0
      on KeyDown: ActivateScreen("1. MAIN", 0)
   Softkey "Softkey_F2" at 0,0 size 0x0
      on KeyDown: ActivateScreen("2. VFD 2 - 5", 0)
   Softkey "Softkey_F3" at 0,0 size 0x0
      on KeyDown: ActivateScreen("3. VFD 6 - 9", 0)
   Softkey "Softkey_F4" at 0,0 size 0x0
      on KeyDown: ActivateScreen("4. VFD 10 - 13", 0)
   Softkey "Softkey_F5" at 0,0 size 0x0
      on KeyDown: ActivateScreen("5. VFD 14 - 17", 0)
   Softkey "Softkey_F6" at 0,0 size 0x0
      on KeyDown: ActivateScreen("6. VFD 18 - 21", 0)
   Softkey "Softkey_F7" at 0,0 size 0x0
      on KeyDown: ActivateScreen("7. VFD 22 - 23", 0)
   Softkey "Softkey_F8" at 0,0 size 0x0
      on KeyDown: ActivateScreen("8. ALARM", 0)
   Softkey "Softkey_F9" at 0,0 size 0x0
      on KeyDown: ActivateScreen("9. VFD PROFIBUS", 0)
   Softkey "Softkey_F10" at 0,0 size 0x0
      on KeyDown: ActivateScreen("10. SETTINGS", 0)

screen "3. VFD 6 - 9" 1280x800, template "Main_Template"
   on GenerateScreen: SetTag("animation_page", 3)
   Bar "Bar_1" at 206,213 size 88x440; MinimumValue 0; MaximumValue 50
      ProcessValue <- "speedActual_address_6"
   Button "Button_7" at 35,514 size 150x62; TextOff '+'
      on Press: function_b14e0dd5("increaseSpeed_address_6", 0)
      Appearance <- "statusIncrease_address_6"
   Button "Button_8" at 35,591 size 150x62; TextOff '-'
      on Press: function_b14e0dd5("decreaseSpeed_address_6", 0)
      Appearance <- "statusDecrease_address_6"
   TextField "Text field_20" at 35,428 size 150x62; Text 'Hz'
   IOField "I/O field_1" at 37,430 size 98x57; FormatPattern 99.99
      ProcessValue <- "speedActual_address_6"
   TextField "Text field_14" at 28,133 size 207x62; Text 'Gauge Roll 1st'
   TextField "Text field_26" at 35,228 size 150x62; Text 'Hz'
   TextField "Text field_32" at 35,328 size 150x62; Text 'Hz'
   IOField "I/O field_2" at 39,231 size 98x57; FormatPattern 99.99
      ProcessValue <- "speedReff_singleSync_address_6"
   TextField "Text field_1" at 35,400 size 115x27; Text 'Actual Speed'
   TextField "Text field_2" at 35,302 size 144x27; Text 'Reff Speed Sync'
   TextField "Text field_3" at 35,200 size 155x27; Text 'Reff Speed Single'
   TextField "Text field_4" at 36,661 size 149x45; Text 'VFD 6'
      Appearance <- "Running_Motor Addres_6"
   Bar "Bar_2" at 518,213 size 88x440; MinimumValue 0; MaximumValue 50
      ProcessValue <- "speedActual_address_7"
   Button "Button_2" at 347,514 size 150x62; TextOff '+'
      on Press: function_b14e0dd5("increaseSpeed_address_7", 0)
      Appearance <- "statusIncrease_address_7"
   Button "Button_3" at 347,591 size 150x62; TextOff '-'
      on Press: function_b14e0dd5("decreaseSpeed_address_7", 0)
      Appearance <- "statusDecrease_address_7"
   TextField "Text field_5" at 347,428 size 150x62; Text 'Hz'
   IOField "I/O field_3" at 349,430 size 98x57; FormatPattern 99.99
      ProcessValue <- "speedActual_address_7"
   TextField "Text field_6" at 340,133 size 207x62; Text 'Conveyor of Gauge Roll 1st'
   TextField "Text field_7" at 347,228 size 150x62; Text 'Hz'
   TextField "Text field_8" at 347,328 size 150x62; Text 'Hz'
   IOField "I/O field_4" at 351,231 size 98x57; FormatPattern 99.99
      ProcessValue <- "speedReff_singleSync_address_7"
   TextField "Text field_9" at 347,400 size 115x27; Text 'Actual Speed'
   TextField "Text field_10" at 347,302 size 144x27; Text 'Reff Speed Sync'
   TextField "Text field_11" at 347,200 size 155x27; Text 'Reff Speed Single'
   TextField "Text field_12" at 348,661 size 149x45; Text 'VFD 7'
      Appearance <- "Running_Motor Addres_7"
   Bar "Bar_3" at 830,213 size 88x440; MinimumValue 0; MaximumValue 50
      ProcessValue <- "speedActual_address_8"
   Button "Button_4" at 659,514 size 150x62; TextOff '+'
      on Press: function_b14e0dd5("increaseSpeed_address_8", 0)
      Appearance <- "statusIncrease_address_8"
   Button "Button_5" at 659,591 size 150x62; TextOff '-'
      on Press: function_b14e0dd5("decreaseSpeed_address_8", 0)
      Appearance <- "statusDecrease_address_8"
   TextField "Text field_13" at 659,428 size 150x62; Text 'Hz'
   IOField "I/O field_5" at 661,430 size 98x57; FormatPattern 99.99
      ProcessValue <- "speedActual_address_8"
   TextField "Text field_15" at 652,133 size 207x62; Text 'Gauge Roll 2nd'
   TextField "Text field_16" at 659,228 size 150x62; Text 'Hz'
   TextField "Text field_17" at 659,328 size 150x62; Text 'Hz'
   IOField "I/O field_6" at 663,231 size 98x57; FormatPattern 99.99
      ProcessValue <- "speedReff_singleSync_address_8"
   TextField "Text field_18" at 659,400 size 115x27; Text 'Actual Speed'
   TextField "Text field_19" at 659,302 size 144x27; Text 'Reff Speed Sync'
   TextField "Text field_21" at 659,200 size 155x27; Text 'Reff Speed Single'
   TextField "Text field_22" at 660,661 size 149x45; Text 'VFD 8'
      Appearance <- "Running_Motor Addres_8"
   Bar "Bar_4" at 1142,213 size 88x440; MinimumValue 0; MaximumValue 50
      ProcessValue <- "speedActual_address_9"
   Button "Button_6" at 971,514 size 150x62; TextOff '+'
      on Press: function_b14e0dd5("increaseSpeed_address_9", 0)
      Appearance <- "statusIncrease_address_9"
   Button "Button_9" at 971,591 size 150x62; TextOff '-'
      on Press: function_b14e0dd5("decreaseSpeed_address_9", 0)
      Appearance <- "statusDecrease_address_9"
   TextField "Text field_23" at 971,428 size 150x62; Text 'Hz'
   IOField "I/O field_7" at 973,430 size 98x57; FormatPattern 99.99
      ProcessValue <- "speedActual_address_9"
   TextField "Text field_24" at 964,133 size 207x62; Text 'Conveyor of Gauge Roll 2nd'
   TextField "Text field_25" at 971,228 size 150x62; Text 'Hz'
   TextField "Text field_27" at 971,328 size 150x62; Text 'Hz'
   IOField "I/O field_8" at 975,231 size 98x57; FormatPattern 99.99
      ProcessValue <- "speedReff_singleSync_address_9"
   TextField "Text field_28" at 971,400 size 115x27; Text 'Actual Speed'
   TextField "Text field_29" at 971,302 size 144x27; Text 'Reff Speed Sync'
   TextField "Text field_30" at 971,200 size 155x27; Text 'Reff Speed Single'
   TextField "Text field_31" at 972,661 size 149x45; Text 'VFD 9'
      Appearance <- "Running_Motor Addres_9"
   IOField "I/O field_14" at 349,330 size 98x57; FormatPattern 99.99
      ProcessValue <- "speedReff_NOT_singleSync_address_7"
   IOField "I/O field_9" at 661,330 size 98x57; FormatPattern 99.99
      ProcessValue <- "speedReff_NOT_singleSync_address_8"
   IOField "I/O field_10" at 973,330 size 98x57; FormatPattern 99.99
      ProcessValue <- "speedReff_NOT_singleSync_address_9"
   SymbolicIOField "Symbolic I/O field_2" at 550,133 size 77x62; TextOn '1'; TextOff '0'; TextList "Mode_Syncron"
      Appearance <- "Syncron_2"
      ProcessValue <- "Syncron_2"
   SymbolicIOField "Symbolic I/O field_3" at 862,133 size 77x62; TextOn '1'; TextOff '0'; TextList "Mode_Syncron"
      Appearance <- "Syncron_2"
      ProcessValue <- "Syncron_2"
   SymbolicIOField "Symbolic I/O field_4" at 1174,133 size 77x62; TextOn '1'; TextOff '0'; TextList "Mode_Syncron"
      Appearance <- "Syncron_2"
      ProcessValue <- "Syncron_2"
   IOField "I/O field_11" at 37,330 size 98x57; FormatPattern 99.99
      ProcessValue <- "speedReff_NOT_singleSync_address_6"
   SymbolicIOField "Symbolic I/O field_1" at 238,133 size 77x62; TextOn '1'; TextOff '0'; TextList "Mode_Syncron"
      Appearance <- "Syncron_2"
      ProcessValue <- "Syncron_2"
   Button "Button_1" at 0,721 size 160x79; TextOff 'MAIN'
      on Click: ActivateScreen("1. MAIN", 0)
      Appearance <- "animation_page"
   Button "Button_10" at 160,721 size 160x79; TextOff 'VFD 2 - 5'
      on Click: ActivateScreen("2. VFD 2 - 5", 0)
      Appearance <- "animation_page"
   Button "Button_11" at 320,721 size 160x79; TextOff 'VFD 6 - 9'
      on Click: ActivateScreen("3. VFD 6 - 9", 0)
      Appearance <- "animation_page"
   Button "Button_12" at 480,721 size 160x79; TextOff 'VFD 10 - 13'
      on Click: ActivateScreen("4. VFD 10 - 13", 0)
      Appearance <- "animation_page"
   Button "Button_13" at 640,721 size 160x79; TextOff 'VFD 14 - 17'
      on Click: ActivateScreen("5. VFD 14 - 17", 0)
      Appearance <- "animation_page"
   Button "Button_14" at 800,721 size 160x79; TextOff 'VFD 18 - 21'
      on Click: ActivateScreen("6. VFD 18 - 21", 0)
      Appearance <- "animation_page"
   Button "Button_15" at 960,721 size 160x79; TextOff 'VFD 22 - 23'
      on Click: ActivateScreen("7. VFD 22 - 23", 0)
      Appearance <- "animation_page"
   Button "Button_16" at 1120,721 size 160x79; TextOff 'Alarm'
      on Click: ActivateScreen("8. ALARM", 0)
      Appearance <- "animation_page"
   TextField "Text field_34" at 0,64 size 331x50; Text 'MOTOR CONTROL SPEED'
   Softkey "Softkey_F1" at 0,0 size 0x0
      on KeyDown: ActivateScreen("1. MAIN", 0)
   Softkey "Softkey_F2" at 0,0 size 0x0
      on KeyDown: ActivateScreen("2. VFD 2 - 5", 0)
   Softkey "Softkey_F3" at 0,0 size 0x0
      on KeyDown: ActivateScreen("3. VFD 6 - 9", 0)
   Softkey "Softkey_F4" at 0,0 size 0x0
      on KeyDown: ActivateScreen("4. VFD 10 - 13", 0)
   Softkey "Softkey_F5" at 0,0 size 0x0
      on KeyDown: ActivateScreen("5. VFD 14 - 17", 0)
   Softkey "Softkey_F6" at 0,0 size 0x0
      on KeyDown: ActivateScreen("6. VFD 18 - 21", 0)
   Softkey "Softkey_F7" at 0,0 size 0x0
      on KeyDown: ActivateScreen("7. VFD 22 - 23", 0)
   Softkey "Softkey_F8" at 0,0 size 0x0
      on KeyDown: ActivateScreen("8. ALARM", 0)
   Softkey "Softkey_F9" at 0,0 size 0x0
      on KeyDown: ActivateScreen("9. VFD PROFIBUS", 0)
   Softkey "Softkey_F10" at 0,0 size 0x0
      on KeyDown: ActivateScreen("10. SETTINGS", 0)